
                   REGION "BUILT TEST STRING"
                       IF #pString >= 1 THEN
                           #lengthTest := CONCAT_WSTRING(IN1 := #_lineBox[#pLineBox],
                                                         IN2 := #space,
                                                         IN3 := #stringBox[#pString]);
                       END_IF;
                   END_REGION

                   REGION "TEST STRING NOT TOO LONG"
                       IF LEN(#lengthTest) <= #maxLength THEN
                           #_lineBox[#pLineBox] := #lengthTest;
                       END_IF;
                   END_REGION

                   REGION "TEST STRING TOO LONG"
                       IF LEN(#lengthTest) > #maxLength THEN
                           #_lineBox[#pLineBox] := "Trim"(#_lineBox[#pLineBox]);
                           #_lineBox[#pLineBox] := "Trim"(#_lineBox[#pLineBox]);
                           #pLineBox := #pLineBox + 1;
                           #_lineBox[#pLineBox] := #stringBox[#pString];
                       END_IF;
                   END_REGION

               END_IF;
           END_REGION

       END_FOR;
   END_REGION

   REGION "RETURN"
       #lineBox := #_lineBox;
   END_REGION
END_FUNCTION

FUNCTION "Word Wrap: Concat Lines" : WString   // FC75, SCL
{ S7_Optimized_Access := 'TRUE' }
VERSION : 0.1
   VAR_INPUT
      lineBox : Array[0..#limitLines] of WString["lStringLen"];
   END_VAR
   VAR_TEMP
      pLine : Int;
      ret : WString;
   END_VAR
   VAR CONSTANT
      space : WString := WSTRING#' ';
      blank : WString;
      lineBreak : WString := WSTRING#'$L';
      limitString : Int := 49;
      limitLines : Int := 9;
   END_VAR
BEGIN
   REGION "FOR EACH LINE"
       FOR #pLine := 0 TO #limitLines DO

           REGION "ON END OF LINE LIST"
               IF #lineBox[#pLine] = #space OR #lineBox[#pLine] = #blank THEN
                   EXIT;
               END_IF;
           END_REGION

           REGION "ON FIRST ELEMENT IN LINE LIST"
               IF #pLine = 0 THEN
                   #ret := #lineBox[#pLine];
               END_IF;
           END_REGION

           REGION "CONSTRUCT OUTPUT"
               IF #pLine >= 1 THEN

                   REGION "NO OP ON LINE BREAK CHARACTER"
                       IF #lineBox[#pLine] = #lineBreak THEN
                           ;// no action required
                       END_IF;
                   END_REGION

                   REGION "CONCATINATION"
                       IF #lineBox[#pLine] <> #lineBreak THEN
                           #ret := CONCAT_WSTRING(IN1 := #ret,
                                                  IN2 := #lineBreak,
                                                  IN3 := #lineBox[#pLine]);
                       END_IF;
                   END_REGION

               END_IF;
           END_REGION


       END_FOR;
   END_REGION

   REGION "RETURN"
       #ret := "Trim"(#ret);
       #"Word Wrap: Concat Lines" := #ret;
   END_REGION
END_FUNCTION

// folder: Utilities/Table Navigation

FUNCTION_BLOCK "Table Nav: End of Data Rollover"   // FB11, SCL
{ S7_Optimized_Access := 'TRUE' }
VERSION : 0.1
   VAR_INPUT
      tblData : Variant;
      tblDisp : Variant;
      nullFlag : Int;
      nullCheck : Variant;
      tableNav : "Nav Bar Data: PLC";
   END_VAR
   VAR_IN_OUT
      rowIndices : Variant;
   END_VAR
   VAR_TEMP
      firstNullIndex : DInt;
      len : Struct
         tblData : DInt;
         tblDisp : DInt;
      END_STRUCT;
      nullCheckVals : Array[0..#lenArrs] of DInt;
      offset : DInt;
      pulses : "Nav Bar Data: PLC";
      RET_VAL : Int;
      retRowIndices : Array[0..#lenArrs] of DInt;
   END_VAR
   VAR CONSTANT
      lenArrs : DInt := 999;
   END_VAR
BEGIN
       REGION "DESCRIPTION"
           (*
           Double checks row indicies against data and rolls over on end of data flag.
           *)
       END_REGION

       REGION "COPY TO LOCAL"
           #RET_VAL := MOVE_BLK_VARIANT(SRC := #rowIndices,
                                        COUNT := CountOfElements(#rowIndices),
                                        SRC_INDEX := 0,
                                        DEST_INDEX := 0,
                                        DEST => #retRowIndices);
           #RET_VAL := MOVE_BLK_VARIANT(SRC := #nullCheck,
                                        COUNT := CountOfElements(#nullCheck),
                                        SRC_INDEX := 0,
                                        DEST_INDEX := 0,
                                        DEST => #nullCheckVals);
       END_REGION

       REGION "GET ARRAY PARAMETERS"
           #len.tblData := UDINT_TO_DINT(CountOfElements(#tblData));
           #len.tblDisp := UDINT_TO_DINT(CountOfElements(#tblDisp));
       END_REGION

       REGION "CALCUALTE ROW INDICIES"
           "Table Nav: Calc Row Indices"(lenTblData := #firstNullIndex,
                                         lenTblDisp := #len.tblDisp,
                                         r1 := #retRowIndices[0],
                                         rowIndicies := #retRowIndices);
       END_REGION

       REGION "RETURN ROW INDICIES"
           #RET_VAL := MOVE_BLK_VARIANT(SRC := #retRowIndices,
                                        COUNT := DINT_TO_UDINT(#len.tblDisp),
                                        SRC_INDEX := 0,
                                        DEST_INDEX := 0,
                                        DEST => #rowIndices);
       END_REGION
END_FUNCTION_BLOCK

FUNCTION_BLOCK "Table Nav"   // FB43, SCL
{ S7_Optimized_Access := 'TRUE' }
VERSION : 0.1
   VAR_INPUT
      first_null_index : DInt;   // if you want to roll over before the end of your array, find the first null index and enter it here
      tblData : Variant;   // array to scan
      tblDisp : Variant;   // viewport array
      tableNav : "Nav Bar Data: PLC";   // table navigation udt
   END_VAR
   VAR_IN_OUT
      rowIndices : Variant;
   END_VAR
   VAR
      "inst Pulses: Table Nav" : "Table Nav: Pulses";
      r1 : DInt;
   END_VAR
   VAR_TEMP
      len : Struct
         tblData : DInt;
         tblDisp : DInt;
      END_STRUCT;
      offset : DInt;
      pulses : "Nav Bar Data: PLC";
      RET_VAL : Int;
      ret_row_indices : Array[0..#lenArrs] of DInt;
      ubound : DInt;
   END_VAR
   VAR CONSTANT
      lenArrs : DInt := 999;
   END_VAR
BEGIN
   REGION "DESCRIPTION"
       (*
       The function returns row indicies indicating the visible rows of a larger
       table determined by standard table navigation buttons.
       The function uses the variant data type to handle tables of any size.
       Rollover and rollunder features are built in.
       Row indices must be output to an array of dint (dimension is flexible).
       *)
   END_REGION


   REGION "GET PRESS PULSES"    
       #"inst Pulses: Table Nav"(press := #tableNav,
                                 pulses => #pulses);
   END_REGION


   REGION "RUN ON BUTTON PRESS"
       IF "Table Nav: Run Trigger"(#pulses) THEN

           REGION "GET ARRAY PARAMETERS"
               #len.tblData := UDINT_TO_DINT(CountOfElements(#tblData));
               #len.tblDisp := UDINT_TO_DINT(CountOfElements(#tblDisp));
           END_REGION

           REGION "CALCULATE UPPER BOUND"
               #ubound := #len.tblData;
               IF #first_null_index <= #len.tblData THEN
                   IF #first_null_index > 0 THEN
                       #ubound := #first_null_index;
                   END_IF;
               END_IF;
           END_REGION

           REGION "CALCULATE OFFSET"
               #offset := "Table Nav: Calculate Offset"(pulses := #pulses,
                                                        lenTblData := #ubound,
                                                        lenTblDisp := #len.tblDisp,
                                                        r1 := #r1);
           END_REGION

           REGION "CALCULATE FIRST ROW"
               #r1 := "Table Nav: Get First Row"(table_length := #ubound,
                                                 offset := #offset,
                                                 first_row := #r1);
           END_REGION

           REGION "CALCUALTE ROW INDICIES"
               "Table Nav: Calc Row Indices"(lenTblData := #ubound,
                                             lenTblDisp := #len.tblDisp,
                                             r1 := #r1,
                                             rowIndicies := #ret_row_indices);
           END_REGION

           REGION "RETURN ROW INDICIES"
               #RET_VAL := MOVE_BLK_VARIANT(SRC := #ret_row_indices,
                                            COUNT := DINT_TO_UDINT(#len.tblDisp),
                                            SRC_INDEX := 0,
                                            DEST_INDEX := 0,
                                            DEST => #rowIndices);
           END_REGION

       END_IF;
   END_REGION
END_FUNCTION_BLOCK

FUNCTION_BLOCK "Table Nav: Pulses"   // FB44, SCL
{ S7_Optimized_Access := 'TRUE' }
VERSION : 0.1
   VAR_INPUT
      press : "Nav Bar Data: PLC";
   END_VAR
   VAR_OUTPUT
      pulses : "Nav Bar Data: PLC";
   END_VAR
   VAR
      old : "Nav Bar Data: PLC";
   END_VAR
BEGIN
   REGION "EVALUATION"
       #pulses.top.actuate := #press.top.actuate AND NOT #old.top.actuate;
       #pulses.pageUp.actuate := #press.pageUp.actuate AND NOT #old.pageUp.actuate;
       #pulses.lineUp.actuate := #press.lineUp.actuate AND NOT #old.lineUp.actuate;
       #pulses.lineDown.actuate := #press.lineDown.actuate AND NOT #old.lineDown.actuate;
       #pulses.pageDown.actuate := #press.pageDown.actuate AND NOT #old.pageDown.actuate;
       #pulses.bottom.actuate := #press.bottom.actuate AND NOT #old.bottom.actuate;
   END_REGION

   REGION "CHANGE DETECTION"
       #old.top.actuate := #press.top.actuate;
       #old.pageUp.actuate := #press.pageUp.actuate;
       #old.lineUp.actuate := #press.lineUp.actuate;
       #old.lineDown.actuate := #press.lineDown.actuate;
       #old.pageDown.actuate := #press.pageDown.actuate;
       #old.bottom.actuate := #press.bottom.actuate;
   END_REGION
END_FUNCTION_BLOCK

FUNCTION "Table Nav: Get Null Index" : DInt   // FC14, SCL
{ S7_Optimized_Access := 'TRUE' }
VERSION : 0.1
   VAR_INPUT
      nullFlag : Int;
      nullCheckVals : Array[0.."wipCount"] of DInt;
   END_VAR
   VAR_TEMP
      pNullCheck : DInt;
   END_VAR
BEGIN
   WHILE #nullCheckVals[#pNullCheck] <> #nullFlag AND #pNullCheck <= "wipCount" DO
       #pNullCheck += 1;
   END_WHILE;
   #"Table Nav: Get Null Index" := #pNullCheck;
END_FUNCTION

FUNCTION "Table Nav: Get First Row" : DInt   // FC44, SCL
{ S7_Optimized_Access := 'TRUE' }
VERSION : 0.1
   VAR_INPUT
      first_row : DInt;
      offset : DInt;
      table_length : DInt;
   END_VAR
   VAR_TEMP
      ret : DInt;
   END_VAR
BEGIN
   REGION "DESCRIPTION"
       (*
       The new first row of the table is calculated from the offset. 
       Rollover and rollunder are resolved for the first row.
       *)
   END_REGION

   REGION "COPY TO INTERNAL"
       #ret := #first_row + #offset;
   END_REGION

   REGION "ROLLUNDER"
       IF #ret < 0 THEN
           #ret := #ret + #table_length;
       END_IF;
   END_REGION

   REGION "ROLLOVER"
       IF #ret > #table_length THEN
           #ret := #ret - #table_length;
       END_IF;
   END_REGION

   REGION "OUTPUT"
       #"Table Nav: Get First Row" := #ret;
   END_REGION
END_FUNCTION

FUNCTION "Table Nav: Calculate Offset" : DInt   // FC45, SCL
{ S7_Optimized_Access := 'TRUE' }
VERSION : 0.1
   VAR_INPUT
      lenTblData : DInt;
      lenTblDisp : DInt;
      pulses : "Nav Bar Data: PLC";
      r1 : DInt;
   END_VAR
   VAR_TEMP
      retOffset : DInt;
   END_VAR
   // Ret_Val : offset from table row 1 from button
BEGIN
   REGION "DESCRIPTION"
       (*
       The offset from the first row of the table is calculated based on the button pressed.
       *)
   END_REGION

   REGION "TOP"
       IF #pulses.top.actuate THEN
           #retOffset := -1 * #r1;
       END_IF;
   END_REGION

   REGION "PAGE UP"
       IF #pulses.pageUp.actuate THEN
           #retOffset := -1 * #lenTblDisp;
       END_IF;
   END_REGION

   REGION "LINE UP"
       IF #pulses.lineUp.actuate THEN
           #retOffset := -1;
       END_IF;
   END_REGION

   REGION "LINE DOWN"
       IF #pulses.lineDown.actuate THEN
           #retOffset := 1;
       END_IF;
   END_REGION

   REGION "PAGE DOWN"
       IF #pulses.pageDown.actuate THEN
           #retOffset := #lenTblDisp ;
       END_IF;
   END_REGION

   REGION "BOTTOM"
       IF #pulses.bottom.actuate THEN
           #retOffset := #lenTblData - #lenTblDisp - #r1;
       END_IF;
   END_REGION

   REGION "RETURN"
       #"Table Nav: Calculate Offset" := #retOffset;
   END_REGION
END_FUNCTION

FUNCTION "Table Nav: Calc Row Indices" : Void   // FC46, SCL
{ S7_Optimized_Access := 'TRUE' }
VERSION : 0.1
   VAR_INPUT
      lenTblData : DInt;
      lenTblDisp : DInt;
      r1 : DInt;
   END_VAR
   VAR_IN_OUT
      rowIndicies : Array[0..#lenRetArr] of DInt;
   END_VAR
   VAR_TEMP
      pOutArr : Int;
      calcRowIdx : DInt;
      retRowIndicies : Array[0..#lenRetArr] of DInt;
   END_VAR
   VAR CONSTANT
      lenRetArr : Int := 999;
   END_VAR
BEGIN
   REGION "DESCRIPTION"
       (*
       An array of the row indicies that the table should display is returned.
       Rollover and rollunder are calculated index by index.
       *) 
   END_REGION

   REGION "INITIALIZE OUTPUT"
       FOR #pOutArr := 0 TO #lenRetArr DO
           #rowIndicies[#pOutArr] := 0;
       END_FOR;
   END_REGION

   REGION "CALCULATE INDICIES"
       FOR #pOutArr := 0 TO DINT_TO_INT(#lenTblDisp) DO

           REGION "CALCULATE INDEX"
               #calcRowIdx := #r1 + INT_TO_DINT(#pOutArr);
           END_REGION

           REGION "ROLL UNDER"
               IF #calcRowIdx < 0 THEN
                   #calcRowIdx := #calcRowIdx + #lenTblDisp;
               END_IF;
           END_REGION

           REGION "ROLL OVER"
               IF #calcRowIdx >= #lenTblData THEN
                   #calcRowIdx := #calcRowIdx - #lenTblData;
               END_IF;
           END_REGION

           REGION "SAVE TO ARRAY"
               #retRowIndicies[#pOutArr] := #calcRowIdx;
           END_REGION

       END_FOR;
   END_REGION

   REGION "OUTPUT"
       #rowIndicies := #retRowIndicies;
   END_REGION
END_FUNCTION

FUNCTION "Table Nav: Run Trigger" : Bool   // FC47, SCL
{ S7_Optimized_Access := 'TRUE' }
VERSION : 0.1
   VAR_INPUT
      pulses : "Nav Bar Data: PLC";
   END_VAR
BEGIN
   #"Table Nav: Run Trigger" :=
       #pulses.top.actuate OR
       #pulses.pageUp.actuate OR
       #pulses.lineUp.actuate OR
       #pulses.lineDown.actuate OR
       #pulses.pageDown.actuate OR
       #pulses.bottom.actuate;
END_FUNCTION

// folder: Utilities/Timer

FUNCTION "Timer: Time to WString" : WString   // FC36, SCL
{ S7_Optimized_Access := 'TRUE' }
VERSION : 0.1
   VAR_INPUT
      "Time" : Time;
   END_VAR
   VAR_TEMP
      "Time as DInt" : DInt;
      "Hours 10s Place" : DInt;
      "Hours 1s Place" : DInt;
      "Minutes 10s Place" : DInt;
      "Minutes 1s Place" : DInt;
      "Seconds 10s Place" : DInt;
      "Seconds 1s Place" : DInt;
      "Time Elements" : Array[0..4] of WString;
      Length : Int;
      "String Box" : WString;
      "DInt Box" : DInt;
   END_VAR
   VAR CONSTANT
      "Milliseconds per 10 Hours" : DInt := 36_000_000;
      "Milliseconds per Hour" : DInt := 3_600_000;
      "Milliseconds per 10 Minutes" : DInt := 600_000;
      "Milliseconds per Minute" : DInt := 60_000;
      "Milliseconds per 10 Seconds" : DInt := 10_000;
      "Milliseconds per Second" : DInt := 1_000;
   END_VAR
BEGIN
   REGION GET INPUT
       #"Time as DInt" := #Time;
   END_REGION

   REGION CONVERT TIME INTO INDIVIDUAL PLACE VALUES
       #"Minutes 10s Place" := #"Time as DInt" / #"Milliseconds per 10 Minutes";
       #"Minutes 1s Place" := (#"Time as DInt" / #"Milliseconds per Minute") MOD 10;
       #"Seconds 10s Place" := (#"Time as DInt" MOD #"Milliseconds per Minute") / #"Milliseconds per 10 Seconds";
       #"Seconds 1s Place" := (#"Time as DInt" / #"Milliseconds per Second") MOD 10;
   END_REGION

   REGION "ADD SIGN"
       #"Time Elements"[0] := wstring#'';
       IF #"Minutes 10s Place" < 0 OR
           #"Minutes 1s Place" < 0 OR
           #"Seconds 10s Place" < 0 OR
           #"Seconds 1s Place" < 0 THEN
            #"Time Elements"[0] := wstring#'-';
       END_IF;
   END_REGION

   REGION CONVERT PLACE VALUES INTO COMPONENT STRINGS
       // MINUTES
       #"DInt Box" := #"Minutes 10s Place" * 10 + #"Minutes 1s Place";
       #"String Box" := DINT_TO_WSTRING(IN := #"DInt Box");
       #"String Box" := "Strip Sign"("WString":=#"String Box");
       #"String Box" := "Add Leading"("Leading Character" := WCHAR#'0',
                                      "Desired Length" := 2,
                                      "String" := #"String Box");
       #"Time Elements"[1] := #"String Box";
       // COLON
       #"Time Elements"[2] := WSTRING#':';
       // SECONDS
       #"DInt Box" := #"Seconds 10s Place" * 10 + #"Seconds 1s Place";
       #"String Box" := DINT_TO_WSTRING(IN := #"DInt Box");
       #"String Box" := "Strip Sign"("WString":=#"String Box");
       #"String Box" := "Add Leading"("Leading Character" := WCHAR#'0',
                                      "Desired Length" := 2,
                                      "String" := #"String Box");
       #"Time Elements"[3] := #"String Box";
   END_REGION


   REGION RETURN VALUE
       #"Timer: Time to WString" := CONCAT_WSTRING(IN1 := #"Time Elements"[0],
                                            IN2 := #"Time Elements"[1],
                                            IN3 := #"Time Elements"[2],
                                            IN4 := #"Time Elements"[3]);
   END_REGION
END_FUNCTION

FUNCTION "Timer: WString to Time" : Time   // FC38, SCL
{ S7_Optimized_Access := 'TRUE' }
VERSION : 0.1
   VAR_INPUT
      WString : WString;
   END_VAR
   VAR_TEMP
      Count : UInt;
      "DInt Box" : DInt;
      "String Box" : WString [5];
      "Time Box" : Time;
      "WChar Array" : Array[0..4] of WChar;
   END_VAR
   VAR CONSTANT
      "ms/(10 hr)" : DInt := 36_000_000;
      "ms/hr" : DInt := 3_600_000;
      "ms/(10 min)" : DInt := 600_000;
      "ms/min" : DInt := 60_000;
      "ms/(10 sec)" : DInt := 10_000;
      "ms/sec" : DInt := 1_000;
   END_VAR
BEGIN
   REGION EXPLODE INPUT

       #"String Box" := #WString;
       IF #"String Box" = WSTRING#'' THEN
           #"String Box" := WSTRING#'00:00';
       END_IF;

       Strg_TO_Chars(Strg := #"String Box",
                     pChars := 0,
                     Cnt => #Count,
                     Chars := #"WChar Array");

   END_REGION

   REGION CONVERT ARRAY ELEMENTS TO TIME

       // 10S OF MINUTES
       #"DInt Box" := WCHAR_TO_DINT(IN := #"WChar Array"[0]) - 16#30;
       #"Time Box" := #"Time Box" + #"DInt Box" * #"ms/(10 min)";

       // MINUTES
       #"DInt Box" := WCHAR_TO_DINT(IN := #"WChar Array"[1]) - 16#30;
       #"Time Box" := #"Time Box" + #"DInt Box" * #"ms/min";

       // 10S OF SECONDS
       #"DInt Box" := WCHAR_TO_DINT(IN := #"WChar Array"[3]) - 16#30;
       #"Time Box" := #"Time Box" + #"DInt Box" * #"ms/(10 sec)";

       // SECONDS
       #"DInt Box" := WCHAR_TO_DINT(IN := #"WChar Array"[4]) - 16#30;
       #"Time Box" := #"Time Box" + #"DInt Box" * #"ms/sec";

   END_REGION


   REGION RETURN VALUE

       #"Timer: WString to Time" := #"Time Box";

   END_REGION
END_FUNCTION

FUNCTION "Timer: WString to Real" : Real   // FC39, SCL
{ S7_Optimized_Access := 'TRUE' }
VERSION : 0.1
   VAR_INPUT
      wstring : WString;
   END_VAR
   VAR CONSTANT
      msPerSec : Real := 1000.0;
   END_VAR
BEGIN
   #"Timer: WString to Real" := DINT_TO_REAL(TIME_TO_DINT("Timer: WString to Time"(#wstring))) / #msPerSec;
END_FUNCTION

FUNCTION "Timer: Real to WString" : WString   // FC40, SCL
{ S7_Optimized_Access := 'TRUE' }
VERSION : 0.1
   VAR_INPUT
      realVal : Real;
   END_VAR
   VAR CONSTANT
      msPerSec : Real := 1000.0;
   END_VAR
BEGIN
   #"Timer: Real to WString" := "Timer: Time to WString"(DINT_TO_TIME(REAL_TO_DINT(#realVal * #msPerSec)));
END_FUNCTION

FUNCTION "Timer" : Void   // FC79, SCL
{ S7_Optimized_Access := 'TRUE' }
VERSION : 0.1
   VAR_INPUT
      delta : Real;
      allotted : Real;
   END_VAR
   VAR_IN_OUT
      elapsed : Real;
      remaining : Real;
   END_VAR
   VAR_TEMP
      _elapsed : Real;
      _remaining : Real;
   END_VAR
BEGIN
   #_elapsed := #elapsed + #delta;
   #_remaining := #allotted - #_elapsed;
   #elapsed := #_elapsed;
   #remaining := #_remaining;
END_FUNCTION

// ===== library types =====

TYPE "PB Data"
   STRUCT
      actuate : Bool;
      animate : USInt;
      enable : Bool;
      label : WString[80];
      listSelect : UInt;
      visible : Bool;
   END_STRUCT;
END_TYPE

TYPE "PB Data: Text Label"
   STRUCT
      actuate : Bool;
      animate : USInt;
      label : WString[20];
   END_STRUCT;
END_TYPE

TYPE "Station Assignment: Button Details Data"
   STRUCT
      alloted : Struct
         animate : USInt;
         value : WString[10];
      END_STRUCT;
      critical : Struct
         animate : USInt;
         value : WString[10];
      END_STRUCT;
      label : Struct
         animate : USInt;
         value : WString[2];
      END_STRUCT;
      partNumber : Struct
         animate : USInt;
         value : WString[40];
      END_STRUCT;
      select : Struct
         actuate : Bool;
         animate : USInt;
      END_STRUCT;
   END_STRUCT;
END_TYPE

TYPE "IO Field Data: Timers"
   STRUCT
      animate : USInt;
      inputFinished : Bool;
      value : WString[5];
   END_STRUCT;
END_TYPE

TYPE "Line Label Data"
   STRUCT
      animate : Struct
         bg : USInt;
         ioField : USInt;
      END_STRUCT;
      inputFinished : Bool;
      value : WString[10];
   END_STRUCT;
END_TYPE

TYPE "Drop Zone Data"
   STRUCT
      animate : Struct
         bg : USInt;
         ioField : USInt;
      END_STRUCT;
      inputFinished : Bool;
      value : WString[10];
   END_STRUCT;
END_TYPE

TYPE "Station Sim Data"
   STRUCT
      stn : Struct
         animate : USInt;
         label : WString[20];
      END_STRUCT;
      btn : Struct
         actuate : Byte;
         animate : Array[0..7] of USInt;
         labels : Array[0..7] of WString [4];
      END_STRUCT;
   END_STRUCT;
END_TYPE

// folder: Main HMI

TYPE "Table Row Data"
   STRUCT
      address : DInt := -1;
      ordered : Bool;
      pbSelection : Struct
         actuate : Bool;
         animate : USInt;
      END_STRUCT;
      rtBackground : Struct
         animate : USInt;
      END_STRUCT;
      tfDropZone : Struct
         animate : USInt;
         value : WString[20];
      END_STRUCT;
      tfLine : Struct
         animate : USInt;
         value : WString[20];
      END_STRUCT;
      tfPartNumber : Struct
         animateDL : USInt;
         animateSL : USInt;
         value : WString[40];
      END_STRUCT;
      tfTime : Struct
         animate : USInt;
         value : WString[20];
      END_STRUCT;
   END_STRUCT;
END_TYPE

(* ===== HMI "HMI_RT_1" =====
system functions are stored by id; their names below are inferred from use
connection "Main HMI": ETHERNET, S7_1500_OMS

HMI tags "Default tag table"
   "Clock_Byte" : Byte = PLC Clock_Byte AT %MB0, 100 ms
   "HMI Data: Warehouse HMI_screenNumber" : Int = PLC "HMI Data: Warehouse HMI".screenNumber AT %DB1.DBW0, 100 ms
   "HMI Data: Warehouse HMI_barcode" : Barcode Screen = PLC "HMI Data: Warehouse HMI".barcode AT %DB1.DBW0, 100 ms
   "HMI Data: Warehouse HMI_tableNav_top" : Push Button Data = PLC "HMI Data: Warehouse HMI".tableNav.top, 100 ms
   "HMI Data: Warehouse HMI_tableNav_pageUp" : Push Button Data = PLC "HMI Data: Warehouse HMI".tableNav.pageUp, 100 ms
   "HMI Data: Warehouse HMI_tableNav_lineUp" : Push Button Data = PLC "HMI Data: Warehouse HMI".tableNav.lineUp, 100 ms
   "HMI Data: Warehouse HMI_tableNav_lineDown" : Push Button Data = PLC "HMI Data: Warehouse HMI".tableNav.lineDown, 100 ms
   "HMI Data: Warehouse HMI_tableNav_pageDown" : Push Button Data = PLC "HMI Data: Warehouse HMI".tableNav.pageDown, 100 ms
   "HMI Data: Warehouse HMI_tableNav_bottom" : Push Button Data = PLC "HMI Data: Warehouse HMI".tableNav.bottom, 100 ms
   "HMI Data: Warehouse HMI_networkHealth_pnioDevices{1}" : Push Button Data = PLC "HMI Data: Warehouse HMI".networkHealth.pnioDevices[1], 100 ms
   "HMI Data: Warehouse HMI_networkHealth_pnioDevices{2}" : Push Button Data = PLC "HMI Data: Warehouse HMI".networkHealth.pnioDevices[2], 100 ms
   "HMI Data: Warehouse HMI_networkHealth_pnioDevices{3}" : Push Button Data = PLC "HMI Data: Warehouse HMI".networkHealth.pnioDevices[3], 100 ms
   "HMI Data: Warehouse HMI_networkHealth_pnioDevices{4}" : Push Button Data = PLC "HMI Data: Warehouse HMI".networkHealth.pnioDevices[4], 100 ms
   "HMI Data: Warehouse HMI_networkHealth_pnioDevices{5}" : Push Button Data = PLC "HMI Data: Warehouse HMI".networkHealth.pnioDevices[5], 100 ms
   "HMI Data: Warehouse HMI_networkHealth_pnioDevices{6}" : Push Button Data = PLC "HMI Data: Warehouse HMI".networkHealth.pnioDevices[6], 100 ms
   "HMI Data: Warehouse HMI_networkHealth_pnioDevices{7}" : Push Button Data = PLC "HMI Data: Warehouse HMI".networkHealth.pnioDevices[7], 100 ms
   "HMI Data: Warehouse HMI_networkHealth_pnioDevices{8}" : Push Button Data = PLC "HMI Data: Warehouse HMI".networkHealth.pnioDevices[8], 100 ms
   "HMI Data: Warehouse HMI_networkHealth_pnioDevices{9}" : Push Button Data = PLC "HMI Data: Warehouse HMI".settings.selectStation, 100 ms
   "HMI Data: Warehouse HMI_networkHealth_pnioDevices{10}" : Push Button Data = PLC "HMI Data: Warehouse HMI".networkHealth.pnioDevices[10], 100 ms
   "HMI Data: Warehouse HMI_networkHealth_pnioDevices{11}" : Push Button Data = PLC "HMI Data: Warehouse HMI".networkHealth.pnioDevices[11], 100 ms
   "HMI Data: Warehouse HMI_networkHealth_pnioDevices{12}" : Push Button Data = PLC "HMI Data: Warehouse HMI".networkHealth.pnioDevices[12], 100 ms
   "HMI Data: Warehouse HMI_networkHealth_pnioDevices{13}" : Push Button Data = PLC "HMI Data: Warehouse HMI".networkHealth.pnioDevices[13], 100 ms
   "HMI Data: Warehouse HMI_networkHealth_pnioDevices{16}" : Push Button Data = PLC "HMI Data: Warehouse HMI".networkHealth.pnioDevices[16], 100 ms
   "HMI Data: Warehouse HMI_networkHealth_pnioDevices{14}" : Push Button Data = PLC "HMI Data: Warehouse HMI".networkHealth.pnioDevices[14], 100 ms
   "HMI Data: Warehouse HMI_networkHealth_pnioDevices{15}" : Push Button Data = PLC "HMI Data: Warehouse HMI".networkHealth.pnioDevices[15], 100 ms
   "HMI Data: Warehouse HMI_networkHealth_pnioDevices{17}" : Push Button Data = PLC "HMI Data: Warehouse HMI".networkHealth.pnioDevices[17], 100 ms
   "HMI Data: Warehouse HMI_networkHealth_pnioDevices{18}" : Push Button Data = PLC "HMI Data: Warehouse HMI".networkHealth.pnioDevices[18], 100 ms
   "HMI Data: Warehouse HMI_networkHealth_pnioDevices{19}" : Push Button Data = PLC "HMI Data: Warehouse HMI".networkHealth.pnioDevices[19], 100 ms
   "HMI Data: Warehouse HMI_networkHealth_pnioDevices{20}" : Push Button Data = PLC "HMI Data: Warehouse HMI".networkHealth.pnioDevices[20], 100 ms
   "HMI Data: Warehouse HMI_networkHealth_pnioDevices{21}" : Push Button Data = PLC "HMI Data: Warehouse HMI".networkHealth.pnioDevices[21], 100 ms
   "HMI Data: Warehouse HMI_networkHealth_pnioDevices{22}" : Push Button Data = PLC "HMI Data: Warehouse HMI".networkHealth.pnioDevices[22], 100 ms
   "HMI Data: Warehouse HMI_networkHealth_pnioDevices{31}" : Push Button Data = PLC "HMI Data: Warehouse HMI".networkHealth.pnioDevices[31], 100 ms
   "HMI Data: Warehouse HMI_networkHealth_pnioDevices{32}" : Push Button Data = PLC "HMI Data: Warehouse HMI".networkHealth.pnioDevices[32], 100 ms
   "HMI Data: Warehouse HMI_networkHealth_pnioDevices{29}" : Push Button Data = PLC "HMI Data: Warehouse HMI".networkHealth.pnioDevices[29], 100 ms
   "HMI Data: Warehouse HMI_networkHealth_pnioDevices{30}" : Push Button Data = PLC "HMI Data: Warehouse HMI".networkHealth.pnioDevices[30], 100 ms
   "HMI Data: Warehouse HMI_networkHealth_pnioDevices{27}" : Push Button Data = PLC "HMI Data: Warehouse HMI".networkHealth.pnioDevices[27], 100 ms
   "HMI Data: Warehouse HMI_networkHealth_pnioDevices{28}" : Push Button Data = PLC "HMI Data: Warehouse HMI".networkHealth.pnioDevices[28], 100 ms
   "HMI Data: Warehouse HMI_networkHealth_pnioDevices{23}" : Push Button Data = PLC "HMI Data: Warehouse HMI".networkHealth.pnioDevices[23], 100 ms
   "HMI Data: Warehouse HMI_networkHealth_pnioDevices{24}" : Push Button Data = PLC "HMI Data: Warehouse HMI".networkHealth.pnioDevices[24], 100 ms
   "HMI Data: Warehouse HMI_networkHealth_pnioDevices{25}" : Push Button Data = PLC "HMI Data: Warehouse HMI".networkHealth.pnioDevices[25], 100 ms
   "HMI Data: Warehouse HMI_networkHealth_pnioDevices{26}" : Push Button Data = PLC "HMI Data: Warehouse HMI".networkHealth.pnioDevices[26], 100 ms
   "HMI Data: Warehouse HMI_networkHealth_pnioDevices{33}" : Push Button Data = PLC "HMI Data: Warehouse HMI".networkHealth.pnioDevices[33], 100 ms
   "HMI Data: Warehouse HMI_networkHealth_pnioDevices{34}" : Push Button Data = PLC "HMI Data: Warehouse HMI".networkHealth.pnioDevices[34], 100 ms
   "HMI Data: Warehouse HMI_networkHealth_pnioDevices{35}" : Push Button Data = PLC "HMI Data: Warehouse HMI".networkHealth.pnioDevices[35], 100 ms
   "HMI Data: Warehouse HMI_networkHealth_pnioDevices{36}" : Push Button Data = PLC "HMI Data: Warehouse HMI".networkHealth.pnioDevices[36], 100 ms
   "HMI Data: Warehouse HMI_networkHealth_pnioDevices{37}" : Push Button Data = PLC "HMI Data: Warehouse HMI".networkHealth.pnioDevices[37], 100 ms
   "HMI Data: Warehouse HMI_networkHealth_pnioDevices{38}" : Push Button Data = PLC "HMI Data: Warehouse HMI".networkHealth.pnioDevices[38], 100 ms
   "HMI Data: Warehouse HMI_networkHealth_pnioDevices{39}" : Push Button Data = PLC "HMI Data: Warehouse HMI".networkHealth.pnioDevices[39], 100 ms
   "HMI Data: Warehouse HMI_networkHealth_pnioDevices{40}" : Push Button Data = PLC "HMI Data: Warehouse HMI".networkHealth.pnioDevices[40], 100 ms
   "HMI Data: Warehouse HMI_networkHealth_pnioDevices{41}" : Push Button Data = PLC "HMI Data: Warehouse HMI".networkHealth.pnioDevices[41], 100 ms
   "HMI Data: Warehouse HMI_networkHealth_pnioDevices{42}" : Push Button Data = PLC "HMI Data: Warehouse HMI".networkHealth.pnioDevices[42], 100 ms
   "HMI Data: Warehouse HMI_networkHealth_pnioDevices{43}" : Push Button Data = PLC "HMI Data: Warehouse HMI".networkHealth.pnioDevices[43], 100 ms
   "HMI Data: Warehouse HMI_networkHealth_pnioDevices{44}" : Push Button Data = PLC "HMI Data: Warehouse HMI".networkHealth.pnioDevices[44], 100 ms
   "HMI Data: Warehouse HMI_networkHealth_pnioDevices{45}" : Push Button Data = PLC "HMI Data: Warehouse HMI".networkHealth.pnioDevices[45], 100 ms
   "HMI Data: Warehouse HMI_networkHealth_pnioDevices{46}" : Push Button Data = PLC "HMI Data: Warehouse HMI".networkHealth.pnioDevices[46], 100 ms
   "HMI Data: Warehouse HMI_networkHealth_pnioDevices{47}" : Push Button Data = PLC "HMI Data: Warehouse HMI".networkHealth.pnioDevices[47], 100 ms
   "HMI Data: Warehouse HMI_networkHealth_pnioDevices{48}" : Push Button Data = PLC "HMI Data: Warehouse HMI".networkHealth.pnioDevices[48], 100 ms
   "HMI Data: Warehouse HMI_networkHealth_et200spPopUp" : Station: ET200SP Comm Debug Data = PLC "HMI Data: Warehouse HMI".networkHealth.et200spPopUp, 100 ms
   "HMI Data: Warehouse HMI_networkHealth_kp8PopUp" : Station: KP8 Comm Debug Data = PLC "HMI Data: Warehouse HMI".networkHealth.kp8PopUp, 100 ms
   "HMI Data: Warehouse HMI_networkHealth_selectedDevice" : Int = PLC "HMI Data: Warehouse HMI".networkHealth.selectedDevice, 100 ms

HMI tags "Pop Ups: Select Buttons"
   "HMI Data: Warehouse HMI_pop_up_select_buttons_buttons{0}" : Push Button Data = PLC "HMI Data: Warehouse HMI".pop_up.select_buttons.buttons[0], 100 ms
   "HMI Data: Warehouse HMI_pop_up_select_buttons_buttons{1}" : Push Button Data = PLC "HMI Data: Warehouse HMI".pop_up.select_buttons.buttons[1], 100 ms
   "HMI Data: Warehouse HMI_pop_up_select_buttons_buttons{2}" : Push Button Data = PLC "HMI Data: Warehouse HMI".pop_up.select_buttons.buttons[2], 100 ms
   "HMI Data: Warehouse HMI_pop_up_select_buttons_buttons{3}" : Push Button Data = PLC "HMI Data: Warehouse HMI".pop_up.select_buttons.buttons[3], 100 ms
   "HMI Data: Warehouse HMI_pop_up_select_buttons_buttons{4}" : Push Button Data = PLC "HMI Data: Warehouse HMI".pop_up.select_buttons.buttons[4], 100 ms
   "HMI Data: Warehouse HMI_pop_up_select_buttons_buttons{5}" : Push Button Data = PLC "HMI Data: Warehouse HMI".pop_up.select_buttons.buttons[5], 100 ms
   "HMI Data: Warehouse HMI_pop_up_select_buttons_buttons{6}" : Push Button Data = PLC "HMI Data: Warehouse HMI".pop_up.select_buttons.buttons[6], 100 ms
   "HMI Data: Warehouse HMI_pop_up_select_buttons_buttons{7}" : Push Button Data = PLC "HMI Data: Warehouse HMI".pop_up.select_buttons.buttons[7], 100 ms
   "HMI Data: Warehouse HMI_pop_up_select_buttons_close_screen" : Push Button Data = PLC "HMI Data: Warehouse HMI".pop_up.select_buttons.close_screen, 100 ms

HMI tags "Pop Ups: Select Stations"
   "HMI Data: Warehouse HMI_pop_up_select_stations_close_screen" : Push Button Data = PLC "HMI Data: Warehouse HMI".pop_up.select_stations.close_screen, 100 ms
   "HMI Data: Warehouse HMI_pop_up_select_stations_nav_bar_hmi" : Nav Bar Data: HMI = PLC "HMI Data: Warehouse HMI".pop_up.select_stations.nav_bar.hmi, 100 ms
   "HMI Data: Warehouse HMI_pop_up_select_stations_stn_select_btns{0}" : Push Button Data = PLC "HMI Data: Warehouse HMI".pop_up.select_stations.stn_select_btns[0], 100 ms
   "HMI Data: Warehouse HMI_pop_up_select_stations_stn_select_btns{1}" : Push Button Data = PLC "HMI Data: Warehouse HMI".pop_up.select_stations.stn_select_btns[1], 100 ms
   "HMI Data: Warehouse HMI_pop_up_select_stations_stn_select_btns{10}" : Push Button Data = PLC "HMI Data: Warehouse HMI".pop_up.select_stations.stn_select_btns[10], 100 ms
   "HMI Data: Warehouse HMI_pop_up_select_stations_stn_select_btns{11}" : Push Button Data = PLC "HMI Data: Warehouse HMI".pop_up.select_stations.stn_select_btns[11], 100 ms
   "HMI Data: Warehouse HMI_pop_up_select_stations_stn_select_btns{2}" : Push Button Data = PLC "HMI Data: Warehouse HMI".pop_up.select_stations.stn_select_btns[2], 100 ms
   "HMI Data: Warehouse HMI_pop_up_select_stations_stn_select_btns{3}" : Push Button Data = PLC "HMI Data: Warehouse HMI".pop_up.select_stations.stn_select_btns[3], 100 ms
   "HMI Data: Warehouse HMI_pop_up_select_stations_stn_select_btns{4}" : Push Button Data = PLC "HMI Data: Warehouse HMI".pop_up.select_stations.stn_select_btns[4], 100 ms
   "HMI Data: Warehouse HMI_pop_up_select_stations_stn_select_btns{5}" : Push Button Data = PLC "HMI Data: Warehouse HMI".pop_up.select_stations.stn_select_btns[5], 100 ms
   "HMI Data: Warehouse HMI_pop_up_select_stations_stn_select_btns{6}" : Push Button Data = PLC "HMI Data: Warehouse HMI".pop_up.select_stations.stn_select_btns[6], 100 ms
   "HMI Data: Warehouse HMI_pop_up_select_stations_stn_select_btns{7}" : Push Button Data = PLC "HMI Data: Warehouse HMI".pop_up.select_stations.stn_select_btns[7], 100 ms
   "HMI Data: Warehouse HMI_pop_up_select_stations_stn_select_btns{8}" : Push Button Data = PLC "HMI Data: Warehouse HMI".pop_up.select_stations.stn_select_btns[8], 100 ms
   "HMI Data: Warehouse HMI_pop_up_select_stations_stn_select_btns{9}" : Push Button Data = PLC "HMI Data: Warehouse HMI".pop_up.select_stations.stn_select_btns[9], 100 ms

HMI tags "Pop Ups: Select WIPs"
   "HMI Data: Warehouse HMI_pop_up_select_WIPs_select_wip_buttons{0}" : Push Button Data = PLC "HMI Data: Warehouse HMI".pop_up.select_WIPs.select_wip_buttons[0], 100 ms
   "HMI Data: Warehouse HMI_pop_up_select_WIPs_select_wip_buttons{1}" : Push Button Data = PLC "HMI Data: Warehouse HMI".pop_up.select_WIPs.select_wip_buttons[1], 100 ms
   "HMI Data: Warehouse HMI_pop_up_select_WIPs_select_wip_buttons{2}" : Push Button Data = PLC "HMI Data: Warehouse HMI".pop_up.select_WIPs.select_wip_buttons[2], 100 ms
   "HMI Data: Warehouse HMI_pop_up_select_WIPs_select_wip_buttons{3}" : Push Button Data = PLC "HMI Data: Warehouse HMI".pop_up.select_WIPs.select_wip_buttons[3], 100 ms
   "HMI Data: Warehouse HMI_pop_up_select_WIPs_select_wip_buttons{4}" : Push Button Data = PLC "HMI Data: Warehouse HMI".pop_up.select_WIPs.select_wip_buttons[4], 100 ms
   "HMI Data: Warehouse HMI_pop_up_select_WIPs_select_wip_buttons{5}" : Push Button Data = PLC "HMI Data: Warehouse HMI".pop_up.select_WIPs.select_wip_buttons[5], 100 ms
   "HMI Data: Warehouse HMI_pop_up_select_WIPs_select_wip_buttons{6}" : Push Button Data = PLC "HMI Data: Warehouse HMI".pop_up.select_WIPs.select_wip_buttons[6], 100 ms
   "HMI Data: Warehouse HMI_pop_up_select_WIPs_close_screen" : Push Button Data = PLC "HMI Data: Warehouse HMI".pop_up.select_WIPs.close_screen, 100 ms
   "HMI Data: Warehouse HMI_pop_up_select_WIPs_nav_bar_hmi" : Nav Bar Data: HMI = PLC "HMI Data: Warehouse HMI".pop_up.select_WIPs.nav_bar.hmi, 100 ms

HMI tags "Part Call"
   "HMI Data: Warehouse HMI_partCall_row{0}" : Table Row = PLC "HMI Data: Warehouse HMI".partCall.row[0], 100 ms
   "HMI Data: Warehouse HMI_partCall_row{1}" : Table Row = PLC "HMI Data: Warehouse HMI".partCall.row[1], 100 ms
   "HMI Data: Warehouse HMI_partCall_row{10}" : Table Row = PLC "HMI Data: Warehouse HMI".partCall.row[10], 100 ms
   "HMI Data: Warehouse HMI_partCall_row{2}" : Table Row = PLC "HMI Data: Warehouse HMI".partCall.row[2], 100 ms
   "HMI Data: Warehouse HMI_partCall_row{3}" : Table Row = PLC "HMI Data: Warehouse HMI".partCall.row[3], 100 ms
   "HMI Data: Warehouse HMI_partCall_row{4}" : Table Row = PLC "HMI Data: Warehouse HMI".partCall.row[4], 100 ms
   "HMI Data: Warehouse HMI_partCall_row{5}" : Table Row = PLC "HMI Data: Warehouse HMI".partCall.row[5], 100 ms
   "HMI Data: Warehouse HMI_partCall_row{6}" : Table Row = PLC "HMI Data: Warehouse HMI".partCall.row[6], 100 ms
   "HMI Data: Warehouse HMI_partCall_row{7}" : Table Row = PLC "HMI Data: Warehouse HMI".partCall.row[7], 100 ms
   "HMI Data: Warehouse HMI_partCall_row{8}" : Table Row = PLC "HMI Data: Warehouse HMI".partCall.row[8], 100 ms
   "HMI Data: Warehouse HMI_partCall_row{9}" : Table Row = PLC "HMI Data: Warehouse HMI".partCall.row[9], 100 ms

HMI tags "Sim Stations"
   "HMI Data: Warehouse HMI_simStations_down" : Push Button Data = PLC "HMI Data: Warehouse HMI".simStations.down, 100 ms
   "HMI Data: Warehouse HMI_simStations_me{0}" : Station: Sim Data = PLC "HMI Data: Warehouse HMI".simStations.me[0] AT %DB1.DBX0.0, 100 ms
   "HMI Data: Warehouse HMI_simStations_me{1}" : Station: Sim Data = PLC "HMI Data: Warehouse HMI".simStations.me[1], 100 ms
   "HMI Data: Warehouse HMI_simStations_me{10}" : Station: Sim Data = PLC "HMI Data: Warehouse HMI".simStations.me[10], 100 ms
   "HMI Data: Warehouse HMI_simStations_me{11}" : Station: Sim Data = PLC "HMI Data: Warehouse HMI".simStations.me[11], 100 ms
   "HMI Data: Warehouse HMI_simStations_me{2}" : Station: Sim Data = PLC "HMI Data: Warehouse HMI".simStations.me[2], 100 ms
   "HMI Data: Warehouse HMI_simStations_me{3}" : Station: Sim Data = PLC "HMI Data: Warehouse HMI".simStations.me[3], 100 ms
   "HMI Data: Warehouse HMI_simStations_me{4}" : Station: Sim Data = PLC "HMI Data: Warehouse HMI".simStations.me[4], 100 ms
   "HMI Data: Warehouse HMI_simStations_me{5}" : Station: Sim Data = PLC "HMI Data: Warehouse HMI".simStations.me[5], 100 ms
   "HMI Data: Warehouse HMI_simStations_me{6}" : Station: Sim Data = PLC "HMI Data: Warehouse HMI".simStations.me[6], 100 ms
   "HMI Data: Warehouse HMI_simStations_me{7}" : Station: Sim Data = PLC "HMI Data: Warehouse HMI".simStations.me[7], 100 ms
   "HMI Data: Warehouse HMI_simStations_me{8}" : Station: Sim Data = PLC "HMI Data: Warehouse HMI".simStations.me[8], 100 ms
   "HMI Data: Warehouse HMI_simStations_me{9}" : Station: Sim Data = PLC "HMI Data: Warehouse HMI".simStations.me[9], 100 ms
   "HMI Data: Warehouse HMI_simStations_up" : Push Button Data = PLC "HMI Data: Warehouse HMI".simStations.up, 100 ms

HMI tags "Settings: Interface"
   "HMI Data: Warehouse HMI_settings_assign" : Push Button Data = PLC "HMI Data: Warehouse HMI".settings.assign, 100 ms
   "HMI Data: Warehouse HMI_settings_partNumber" : IO Field Data: Label with Data = PLC "HMI Data: Warehouse HMI".settings.partNumber, 100 ms
   "HMI Data: Warehouse HMI_settings_critical" : IO Field Data: Label with Data = PLC "HMI Data: Warehouse HMI".settings.critical, 100 ms
   "HMI Data: Warehouse HMI_settings_total" : IO Field Data: Label with Data = PLC "HMI Data: Warehouse HMI".settings.total, 100 ms
   "HMI Data: Warehouse HMI_settings_dropzone" : IO Field Data: Label with Data = PLC "HMI Data: Warehouse HMI".settings.dropzone, 100 ms
   "HMI Data: Warehouse HMI_settings_line" : IO Field Data: Label with Data = PLC "HMI Data: Warehouse HMI".settings.line, 100 ms
   "HMI Data: Warehouse HMI_settings_selectButton" : Push Button Data = PLC "HMI Data: Warehouse HMI".settings.selectButton, 100 ms
   "HMI Data: Warehouse HMI_settings_selectWip" : Push Button Data = PLC "HMI Data: Warehouse HMI".settings.selectWip, 100 ms
   "HMI Data: Warehouse HMI_settings_selectStation" : Push Button Data = PLC "HMI Data: Warehouse HMI".settings.selectStation, 100 ms
   "HMI Data: Warehouse HMI_settings_stnTableNavBar_hmi" : Nav Bar Data: HMI = PLC "HMI Data: Warehouse HMI".settings.stnTableNavBar.hmi AT %DB1.DBW0, 100 ms

HMI tags "Settings: Feedback"
   "HMI Data: Warehouse HMI_settings_stationRows{0}" : Settings Station Row Data = PLC "HMI Data: Warehouse HMI".settings.stationRows[0], 100 ms
   "HMI Data: Warehouse HMI_settings_stationRows{1}" : Settings Station Row Data = PLC "HMI Data: Warehouse HMI".settings.stationRows[1], 100 ms
   "HMI Data: Warehouse HMI_settings_stationRows{2}" : Settings Station Row Data = PLC "HMI Data: Warehouse HMI".settings.stationRows[2], 100 ms

graphic list "Vertical Table Nav Bar": 0 '100 x 100 Top'; 1 '100 x 100 Actuated Top'; 2 '100 x 100 Page Up'; 3 '100 x 100 Actuated Page Up'; 4 '100 x 100 Line Up'; 5 '100 x 100 Actuated Line Up'; 6 '100 x 100 Line Down'; 7 '100 x 100 Actuated Line Down'; 8 '100 x 100 Page Down'; 9 '100 x 100 Actuated Page Down'; 10 '100 x 100 Bottom'; 11 '100 x 100 Actuated Bottom'

screen "1 PART CALL" 1366x768
   on GenerateScreen: SetTag("HMI Data: Warehouse HMI_screenNumber", 1)
   Rectangle "Settings Tab Background" at 682,0 size 684x68
      Appearance <- "HMI Data: Warehouse HMI_screenNumber"
   Rectangle "Part Call Tab Background" at 0,0 size 685x68
      Appearance <- "HMI Data: Warehouse HMI_screenNumber"
   Rectangle "Settings Tab Border Hide" at 685,61 size 678x20
      Visibility <- "HMI Data: Warehouse HMI_screenNumber"
   Rectangle "Part Call Tab Border Hide" at 3,61 size 679x20
      Visibility <- "HMI Data: Warehouse HMI_screenNumber"
   Button "Settings Screen" at 683,0 size 683x68; TextOff 'SETTINGS'; Authorization "User administration"
      on Release: ActivateScreen("2 SETTINGS", 0)
   Button "Part Call Screen" at 0,0 size 683x68; TextOff 'PART CALL'
      on Release: ActivateScreen("1 PART CALL", 0)
   TextField "Header Line" at 32,112 size 216x53; Text 'LINE'
   TextField "Header Drop Zone" at 238,112 size 236x53; Text 'DROP ZONE'
   TextField "Header Part Number" at 474,112 size 648x53; Text 'PART NUMBER'
   TextField "Header Time" at 1112,112 size 222x53; Text 'TIME'
   ScreenModuleView "TableRow00" at 27,170 size 1312x52; ScreenModuleType ""
      Guid_{11997190-27688} <- "HMI Data: Warehouse HMI_partCall_row{0}"
      on Guid_{11997190-83214}: ActivateScreen("3 BARCODE", 0)
   ScreenModuleView "TableRow01" at 27,222 size 1312x52; ScreenModuleType ""
      Guid_{11997190-27688} <- "HMI Data: Warehouse HMI_partCall_row{1}"
      on Guid_{11997190-83214}: ActivateScreen("3 BARCODE", 0)
   ScreenModuleView "TableRow02" at 27,274 size 1312x52; ScreenModuleType ""
      Guid_{11997190-27688} <- "HMI Data: Warehouse HMI_partCall_row{2}"
      on Guid_{11997190-83214}: ActivateScreen("3 BARCODE", 0)
   ScreenModuleView "TableRow03" at 27,326 size 1312x52; ScreenModuleType ""
      Guid_{11997190-27688} <- "HMI Data: Warehouse HMI_partCall_row{3}"
      on Guid_{11997190-83214}: ActivateScreen("3 BARCODE", 0)
   ScreenModuleView "TableRow04" at 27,378 size 1312x52; ScreenModuleType ""
      Guid_{11997190-27688} <- "HMI Data: Warehouse HMI_partCall_row{4}"
      on Guid_{11997190-83214}: ActivateScreen("3 BARCODE", 0)
   ScreenModuleView "TableRow05" at 27,430 size 1312x52; ScreenModuleType ""
      Guid_{11997190-27688} <- "HMI Data: Warehouse HMI_partCall_row{5}"
      on Guid_{11997190-83214}: ActivateScreen("3 BARCODE", 0)
   ScreenModuleView "TableRow06" at 27,482 size 1312x52; ScreenModuleType ""
      Guid_{11997190-27688} <- "HMI Data: Warehouse HMI_partCall_row{6}"
      on Guid_{11997190-83214}: ActivateScreen("3 BARCODE", 0)
   ScreenModuleView "TableRow07" at 27,534 size 1312x52; ScreenModuleType ""
      Guid_{11997190-27688} <- "HMI Data: Warehouse HMI_partCall_row{7}"
      on Guid_{11997190-83214}: ActivateScreen("3 BARCODE", 0)
   ScreenModuleView "TableRow08" at 27,586 size 1312x52; ScreenModuleType ""
      Guid_{11997190-27688} <- "HMI Data: Warehouse HMI_partCall_row{8}"
      on Guid_{11997190-83214}: ActivateScreen("3 BARCODE", 0)
   ScreenModuleView "TableRow09" at 27,638 size 1312x52; ScreenModuleType ""
      Guid_{11997190-27688} <- "HMI Data: Warehouse HMI_partCall_row{9}"
      on Guid_{11997190-83214}: ActivateScreen("3 BARCODE", 0)
   ScreenModuleView "TableRow10" at 27,690 size 1312x52; ScreenModuleType ""
      Guid_{11997190-27688} <- "HMI Data: Warehouse HMI_partCall_row{10}"
      on Guid_{11997190-83214}: ActivateScreen("3 BARCODE", 0)

SlideinScreen "GraphX_Slidein_Bottom" 1366x80
   ScreenModuleView "Top" at 0,0 size 227x80; Guid_{11997190-63799} "Top"; ScreenModuleType ""
      Guid_{11997190-63779} <- "HMI Data: Warehouse HMI_tableNav_top"
   ScreenModuleView "Page Up" at 227,0 size 228x80; Guid_{11997190-63799} "pageUp"; ScreenModuleType ""
      Guid_{11997190-63779} <- "HMI Data: Warehouse HMI_tableNav_pageUp"
   ScreenModuleView "Line Up" at 455,0 size 228x80; Guid_{11997190-63799} "Up"; ScreenModuleType ""
      Guid_{11997190-63779} <- "HMI Data: Warehouse HMI_tableNav_lineUp"
   ScreenModuleView "Line Down" at 683,0 size 228x80; Guid_{11997190-63799} "Down"; ScreenModuleType ""
      Guid_{11997190-63779} <- "HMI Data: Warehouse HMI_tableNav_lineDown"
   ScreenModuleView "Page Down" at 911,0 size 228x80; Guid_{11997190-63799} "PageDown"; ScreenModuleType ""
      Guid_{11997190-63779} <- "HMI Data: Warehouse HMI_tableNav_pageDown"
   ScreenModuleView "Bottom" at 1138,0 size 228x80; Guid_{11997190-63799} "Bottom"; ScreenModuleType ""
      Guid_{11997190-63779} <- "HMI Data: Warehouse HMI_tableNav_bottom"
   TextField "Text field_1" at 0,0 size 1366x80; Text 'NOT USED'
      Visibility <- "HMI Data: Warehouse HMI_screenNumber"

SlideinScreen "GraphX_Slidein_Right" 449x768
   ScreenModuleView "Station Sim_1" at 5,5 size 106x232; ScreenModuleType ""
      Guid_{11997190-89108} <- "HMI Data: Warehouse HMI_simStations_me{0}"
   ScreenModuleView "Station Sim_2" at 116,5 size 106x232; ScreenModuleType ""
      Guid_{11997190-89108} <- "HMI Data: Warehouse HMI_simStations_me{1}"
   ScreenModuleView "Station Sim_3" at 227,5 size 106x232; ScreenModuleType ""
      Guid_{11997190-89108} <- "HMI Data: Warehouse HMI_simStations_me{2}"
   ScreenModuleView "Station Sim_4" at 338,5 size 106x232; ScreenModuleType ""
      Guid_{11997190-89108} <- "HMI Data: Warehouse HMI_simStations_me{3}"
   ScreenModuleView "Station Sim_5" at 5,242 size 106x232; ScreenModuleType ""
      Guid_{11997190-89108} <- "HMI Data: Warehouse HMI_simStations_me{4}"
   ScreenModuleView "Station Sim_6" at 5,479 size 106x232; ScreenModuleType ""
      Guid_{11997190-89108} <- "HMI Data: Warehouse HMI_simStations_me{8}"
   ScreenModuleView "Station Sim_7" at 116,242 size 106x232; ScreenModuleType ""
      Guid_{11997190-89108} <- "HMI Data: Warehouse HMI_simStations_me{5}"
   ScreenModuleView "Station Sim_8" at 227,242 size 106x232; ScreenModuleType ""
      Guid_{11997190-89108} <- "HMI Data: Warehouse HMI_simStations_me{6}"
   ScreenModuleView "Station Sim_9" at 338,242 size 106x232; ScreenModuleType ""
      Guid_{11997190-89108} <- "HMI Data: Warehouse HMI_simStations_me{7}"
   ScreenModuleView "Station Sim_10" at 116,479 size 106x232; ScreenModuleType ""
      Guid_{11997190-89108} <- "HMI Data: Warehouse HMI_simStations_me{9}"
   ScreenModuleView "Station Sim_11" at 227,478 size 106x232; ScreenModuleType ""
      Guid_{11997190-89108} <- "HMI Data: Warehouse HMI_simStations_me{10}"
   ScreenModuleView "Station Sim_12" at 338,477 size 106x232; ScreenModuleType ""
      Guid_{11997190-89108} <- "HMI Data: Warehouse HMI_simStations_me{11}"
   ScreenModuleView "PB: Graphic/Text List_1" at 5,716 size 65x45; Guid_{11997190-63799} "Up"; ScreenModuleType ""
      Guid_{11997190-63779} <- "HMI Data: Warehouse HMI_simStations_up"
   ScreenModuleView "PB: Graphic/Text List_2" at 379,716 size 65x45; Guid_{11997190-63799} "Down"; ScreenModuleType ""
      Guid_{11997190-63779} <- "HMI Data: Warehouse HMI_simStations_down"

